REGION Network 13: IW824 - Spare Input
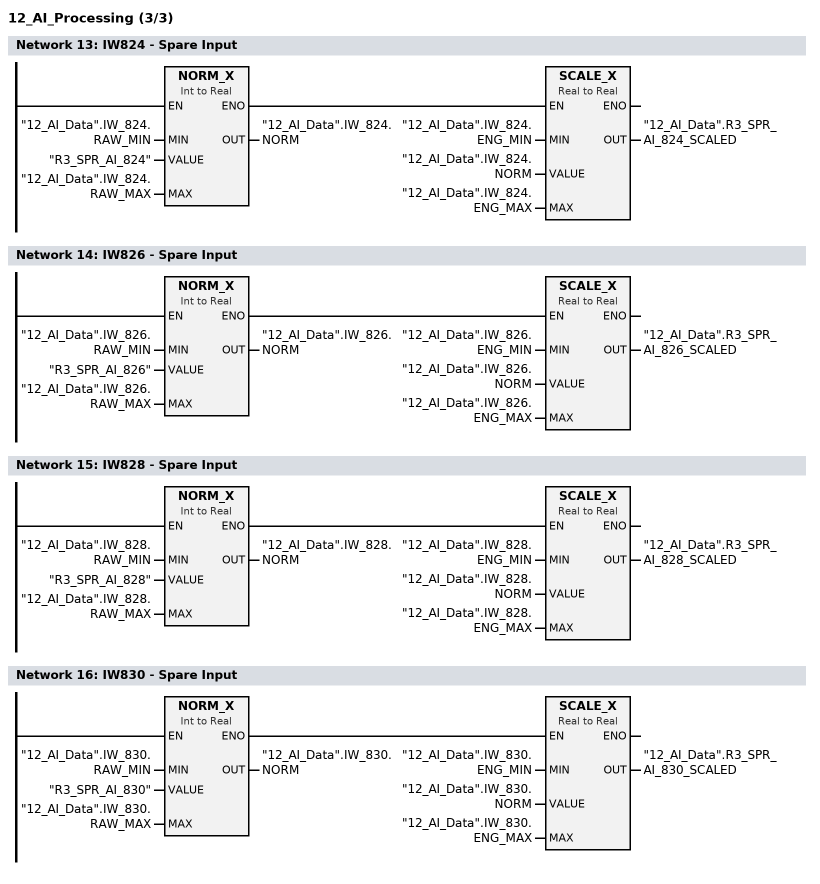
   RUNG wire#powerrail
      { S7_Templates := "[SrcType := Int, DestType := Real]" } Normalize(min := "12_AI_Data".IW_824.RAW_MIN, value := "R3_SPR_AI_824", max := "12_AI_Data".IW_824.RAW_MAX, out => "12_AI_Data".IW_824.NORM)
      { S7_Templates := "[SrcType := Real, DestType := Real]" } Scale(min := "12_AI_Data".IW_824.ENG_MIN, value := "12_AI_Data".IW_824.NORM, max := "12_AI_Data".IW_824.ENG_MAX, out => "12_AI_Data".R3_SPR_AI_824_SCALED)
   END_RUNG
   // the same network as SCL:
   "12_AI_Data".IW_824.NORM := NORM_X(MIN := "12_AI_Data".IW_824.RAW_MIN, VALUE := "R3_SPR_AI_824", MAX := "12_AI_Data".IW_824.RAW_MAX);
   "12_AI_Data".R3_SPR_AI_824_SCALED := SCALE_X(MIN := "12_AI_Data".IW_824.ENG_MIN, VALUE := "12_AI_Data".IW_824.NORM, MAX := "12_AI_Data".IW_824.ENG_MAX);
END_REGION

REGION Network 14: IW826 - Spare Input
   RUNG wire#powerrail
      { S7_Templates := "[SrcType := Int, DestType := Real]" } Normalize(min := "12_AI_Data".IW_826.RAW_MIN, value := "R3_SPR_AI_826", max := "12_AI_Data".IW_826.RAW_MAX, out => "12_AI_Data".IW_826.NORM)
      { S7_Templates := "[SrcType := Real, DestType := Real]" } Scale(min := "12_AI_Data".IW_826.ENG_MIN, value := "12_AI_Data".IW_826.NORM, max := "12_AI_Data".IW_826.ENG_MAX, out => "12_AI_Data".R3_SPR_AI_826_SCALED)
   END_RUNG
   // the same network as SCL:
   "12_AI_Data".IW_826.NORM := NORM_X(MIN := "12_AI_Data".IW_826.RAW_MIN, VALUE := "R3_SPR_AI_826", MAX := "12_AI_Data".IW_826.RAW_MAX);
   "12_AI_Data".R3_SPR_AI_826_SCALED := SCALE_X(MIN := "12_AI_Data".IW_826.ENG_MIN, VALUE := "12_AI_Data".IW_826.NORM, MAX := "12_AI_Data".IW_826.ENG_MAX);
END_REGION

REGION Network 15: IW828 - Spare Input
   RUNG wire#powerrail
      { S7_Templates := "[SrcType := Int, DestType := Real]" } Normalize(min := "12_AI_Data".IW_828.RAW_MIN, value := "R3_SPR_AI_828", max := "12_AI_Data".IW_828.RAW_MAX, out => "12_AI_Data".IW_828.NORM)
      { S7_Templates := "[SrcType := Real, DestType := Real]" } Scale(min := "12_AI_Data".IW_828.ENG_MIN, value := "12_AI_Data".IW_828.NORM, max := "12_AI_Data".IW_828.ENG_MAX, out => "12_AI_Data".R3_SPR_AI_828_SCALED)
   END_RUNG
   // the same network as SCL:
   "12_AI_Data".IW_828.NORM := NORM_X(MIN := "12_AI_Data".IW_828.RAW_MIN, VALUE := "R3_SPR_AI_828", MAX := "12_AI_Data".IW_828.RAW_MAX);
   "12_AI_Data".R3_SPR_AI_828_SCALED := SCALE_X(MIN := "12_AI_Data".IW_828.ENG_MIN, VALUE := "12_AI_Data".IW_828.NORM, MAX := "12_AI_Data".IW_828.ENG_MAX);
END_REGION

REGION Network 16: IW830 - Spare Input
   RUNG wire#powerrail
      { S7_Templates := "[SrcType := Int, DestType := Real]" } Normalize(min := "12_AI_Data".IW_830.RAW_MIN, value := "R3_SPR_AI_830", max := "12_AI_Data".IW_830.RAW_MAX, out => "12_AI_Data".IW_830.NORM)
      { S7_Templates := "[SrcType := Real, DestType := Real]" } Scale(min := "12_AI_Data".IW_830.ENG_MIN, value := "12_AI_Data".IW_830.NORM, max := "12_AI_Data".IW_830.ENG_MAX, out => "12_AI_Data".R3_SPR_AI_830_SCALED)
   END_RUNG
   // the same network as SCL:
   "12_AI_Data".IW_830.NORM := NORM_X(MIN := "12_AI_Data".IW_830.RAW_MIN, VALUE := "R3_SPR_AI_830", MAX := "12_AI_Data".IW_830.RAW_MAX);
   "12_AI_Data".R3_SPR_AI_830_SCALED := SCALE_X(MIN := "12_AI_Data".IW_830.ENG_MIN, VALUE := "12_AI_Data".IW_830.NORM, MAX := "12_AI_Data".IW_830.ENG_MAX);
END_REGION
END_FUNCTION

FUNCTION "14_DQ_Processing" : Void   // FC14, LAD
TITLE = Digital Output Processing
{ S7_Optimized_Access := 'TRUE' }
AUTHOR : JRS
VERSION : 0.1
// To process code outputs prior to physical connection
BEGIN

REGION Network 1: Q136.0 - Fresh Water Fill Valve Control (CV-358)
   // True = OPEN, False = CLOSE
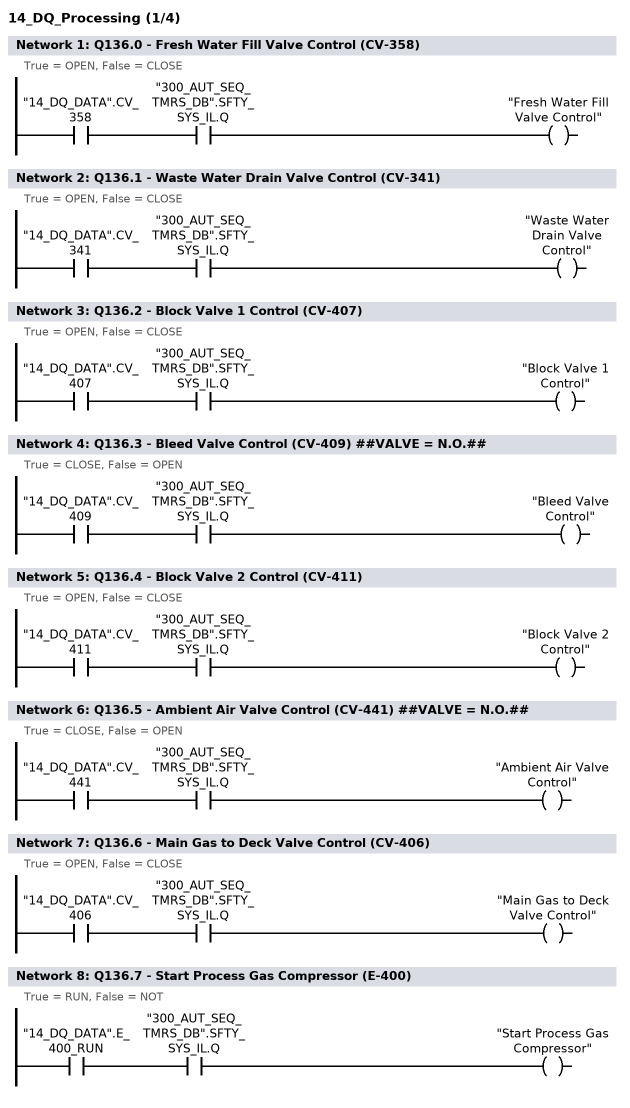
   RUNG wire#powerrail
      Contact( "14_DQ_DATA".CV_358 )
      Contact( "300_AUT_SEQ_TMRS_DB".SFTY_SYS_IL.Q )
      Coil( "Fresh Water Fill Valve Control" )
   END_RUNG
   // the same network as SCL:
   "Fresh Water Fill Valve Control" := "14_DQ_DATA".CV_358 AND "300_AUT_SEQ_TMRS_DB".SFTY_SYS_IL.Q;
END_REGION

REGION Network 2: Q136.1 - Waste Water Drain Valve Control (CV-341)
   // True = OPEN, False = CLOSE
   RUNG wire#powerrail
      Contact( "14_DQ_DATA".CV_341 )
      Contact( "300_AUT_SEQ_TMRS_DB".SFTY_SYS_IL.Q )
      Coil( "Waste Water Drain Valve Control" )
   END_RUNG
   // the same network as SCL:
   "Waste Water Drain Valve Control" := "14_DQ_DATA".CV_341 AND "300_AUT_SEQ_TMRS_DB".SFTY_SYS_IL.Q;
END_REGION

REGION Network 3: Q136.2 - Block Valve 1 Control (CV-407)
   // True = OPEN, False = CLOSE
   RUNG wire#powerrail
      Contact( "14_DQ_DATA".CV_407 )
      Contact( "300_AUT_SEQ_TMRS_DB".SFTY_SYS_IL.Q )
      Coil( "Block Valve 1 Control" )
   END_RUNG
   // the same network as SCL:
   "Block Valve 1 Control" := "14_DQ_DATA".CV_407 AND "300_AUT_SEQ_TMRS_DB".SFTY_SYS_IL.Q;
END_REGION

REGION Network 4: Q136.3 - Bleed Valve Control (CV-409) ##VALVE = N.O.##
   // True = CLOSE, False = OPEN
   RUNG wire#powerrail
      Contact( "14_DQ_DATA".CV_409 )
      Contact( "300_AUT_SEQ_TMRS_DB".SFTY_SYS_IL.Q )
      Coil( "Bleed Valve Control" )
   END_RUNG
   // the same network as SCL:
   "Bleed Valve Control" := "14_DQ_DATA".CV_409 AND "300_AUT_SEQ_TMRS_DB".SFTY_SYS_IL.Q;
END_REGION

REGION Network 5: Q136.4 - Block Valve 2 Control (CV-411)
   // True = OPEN, False = CLOSE
   RUNG wire#powerrail
      Contact( "14_DQ_DATA".CV_411 )
      Contact( "300_AUT_SEQ_TMRS_DB".SFTY_SYS_IL.Q )
      Coil( "Block Valve 2 Control" )
   END_RUNG
   // the same network as SCL:
   "Block Valve 2 Control" := "14_DQ_DATA".CV_411 AND "300_AUT_SEQ_TMRS_DB".SFTY_SYS_IL.Q;
END_REGION

REGION Network 6: Q136.5 - Ambient Air Valve Control (CV-441) ##VALVE = N.O.##
   // True = CLOSE, False = OPEN
   RUNG wire#powerrail
      Contact( "14_DQ_DATA".CV_441 )
      Contact( "300_AUT_SEQ_TMRS_DB".SFTY_SYS_IL.Q )
      Coil( "Ambient Air Valve Control" )
   END_RUNG
   // the same network as SCL:
   "Ambient Air Valve Control" := "14_DQ_DATA".CV_441 AND "300_AUT_SEQ_TMRS_DB".SFTY_SYS_IL.Q;
END_REGION

REGION Network 7: Q136.6 - Main Gas to Deck Valve Control (CV-406)
   // True = OPEN, False = CLOSE
   RUNG wire#powerrail
      Contact( "14_DQ_DATA".CV_406 )
      Contact( "300_AUT_SEQ_TMRS_DB".SFTY_SYS_IL.Q )
      Coil( "Main Gas to Deck Valve Control" )
   END_RUNG
   // the same network as SCL:
   "Main Gas to Deck Valve Control" := "14_DQ_DATA".CV_406 AND "300_AUT_SEQ_TMRS_DB".SFTY_SYS_IL.Q;
END_REGION

REGION Network 8: Q136.7 - Start Process Gas Compressor (E-400)
   // True = RUN, False = NOT
   RUNG wire#powerrail
      Contact( "14_DQ_DATA".E_400_RUN )
      Contact( "300_AUT_SEQ_TMRS_DB".SFTY_SYS_IL.Q )
      Coil( "Start Process Gas Compressor" )
   END_RUNG
   // the same network as SCL:
   "Start Process Gas Compressor" := "14_DQ_DATA".E_400_RUN AND "300_AUT_SEQ_TMRS_DB".SFTY_SYS_IL.Q;
END_REGION

REGION Network 9: Q137.0 - GCU Recirculation Pump Control (P-303)
   // True = RUN, False = NOT
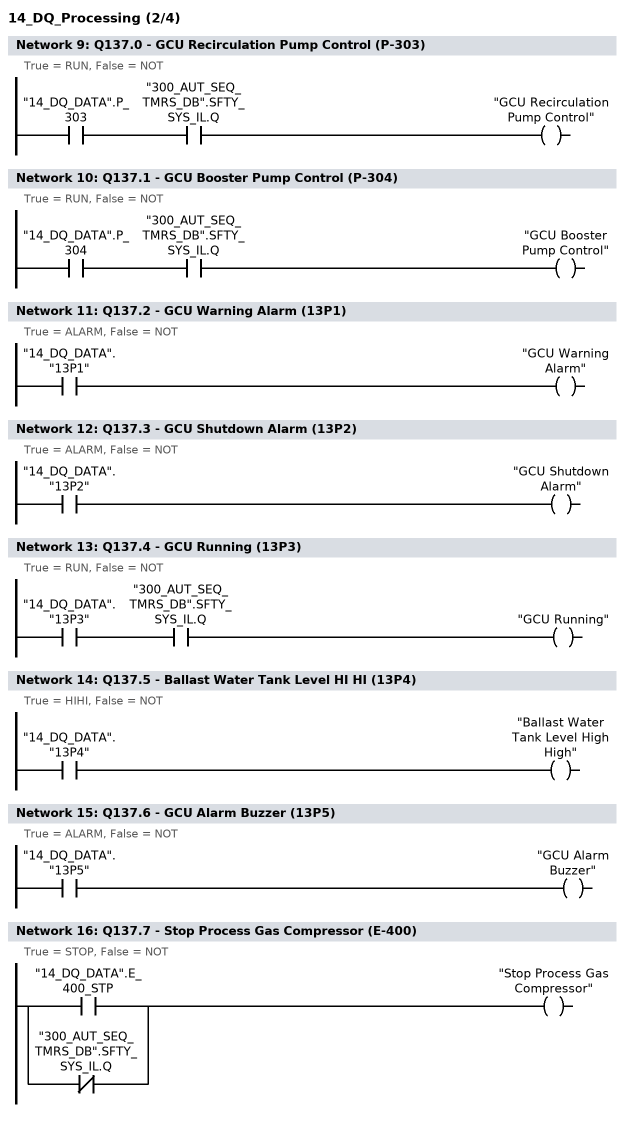
   RUNG wire#powerrail
      Contact( "14_DQ_DATA".P_303 )
      Contact( "300_AUT_SEQ_TMRS_DB".SFTY_SYS_IL.Q )
      Coil( "GCU Recirculation Pump Control" )
   END_RUNG
   // the same network as SCL:
   "GCU Recirculation Pump Control" := "14_DQ_DATA".P_303 AND "300_AUT_SEQ_TMRS_DB".SFTY_SYS_IL.Q;
END_REGION

REGION Network 10: Q137.1 - GCU Booster Pump Control (P-304)
   // True = RUN, False = NOT
   RUNG wire#powerrail
      Contact( "14_DQ_DATA".P_304 )
      Contact( "300_AUT_SEQ_TMRS_DB".SFTY_SYS_IL.Q )
      Coil( "GCU Booster Pump Control" )
   END_RUNG
   // the same network as SCL:
   "GCU Booster Pump Control" := "14_DQ_DATA".P_304 AND "300_AUT_SEQ_TMRS_DB".SFTY_SYS_IL.Q;
END_REGION

REGION Network 11: Q137.2 - GCU Warning Alarm (13P1)
   // True = ALARM, False = NOT
   RUNG wire#powerrail
      Contact( "14_DQ_DATA"."13P1" )
      Coil( "GCU Warning Alarm" )
   END_RUNG
   // the same network as SCL:
   "GCU Warning Alarm" := "14_DQ_DATA"."13P1";
END_REGION

REGION Network 12: Q137.3 - GCU Shutdown Alarm (13P2)
   // True = ALARM, False = NOT
   RUNG wire#powerrail
      Contact( "14_DQ_DATA"."13P2" )
      Coil( "GCU Shutdown Alarm" )
   END_RUNG
   // the same network as SCL:
   "GCU Shutdown Alarm" := "14_DQ_DATA"."13P2";
END_REGION

REGION Network 13: Q137.4 - GCU Running (13P3)
   // True = RUN, False = NOT
   RUNG wire#powerrail
      Contact( "14_DQ_DATA"."13P3" )
      Contact( "300_AUT_SEQ_TMRS_DB".SFTY_SYS_IL.Q )
      Coil( "GCU Running" )
   END_RUNG
   // the same network as SCL:
   "GCU Running" := "14_DQ_DATA"."13P3" AND "300_AUT_SEQ_TMRS_DB".SFTY_SYS_IL.Q;
END_REGION

REGION Network 14: Q137.5 - Ballast Water Tank Level HI HI (13P4)
   // True = HIHI, False = NOT
   RUNG wire#powerrail
      Contact( "14_DQ_DATA"."13P4" )
      Coil( "Ballast Water Tank Level High High" )
   END_RUNG
   // the same network as SCL:
   "Ballast Water Tank Level High High" := "14_DQ_DATA"."13P4";
END_REGION

REGION Network 15: Q137.6 - GCU Alarm Buzzer (13P5)
   // True = ALARM, False = NOT
   RUNG wire#powerrail
      Contact( "14_DQ_DATA"."13P5" )
      Coil( "GCU Alarm Buzzer" )
   END_RUNG
   // the same network as SCL:
   "GCU Alarm Buzzer" := "14_DQ_DATA"."13P5";
END_REGION

REGION Network 16: Q137.7 - Stop Process Gas Compressor (E-400)
   // True = STOP, False = NOT
   RUNG wire#powerrail
      Contact( "14_DQ_DATA".E_400_STP )
      wire#w1
      Coil( "Stop Process Gas Compressor" )
   END_RUNG
   RUNG wire#powerrail
      I_Contact( "300_AUT_SEQ_TMRS_DB".SFTY_SYS_IL.Q )
   END_RUNG wire#w1
   // the same network as SCL:
   "Stop Process Gas Compressor" := "14_DQ_DATA".E_400_STP OR NOT "300_AUT_SEQ_TMRS_DB".SFTY_SYS_IL.Q;
END_REGION

REGION Network 17: Q138.0 - Pilot For GTT FPT Valve (CV-422-FPT)
   // True = OPEN, False = CLOSE
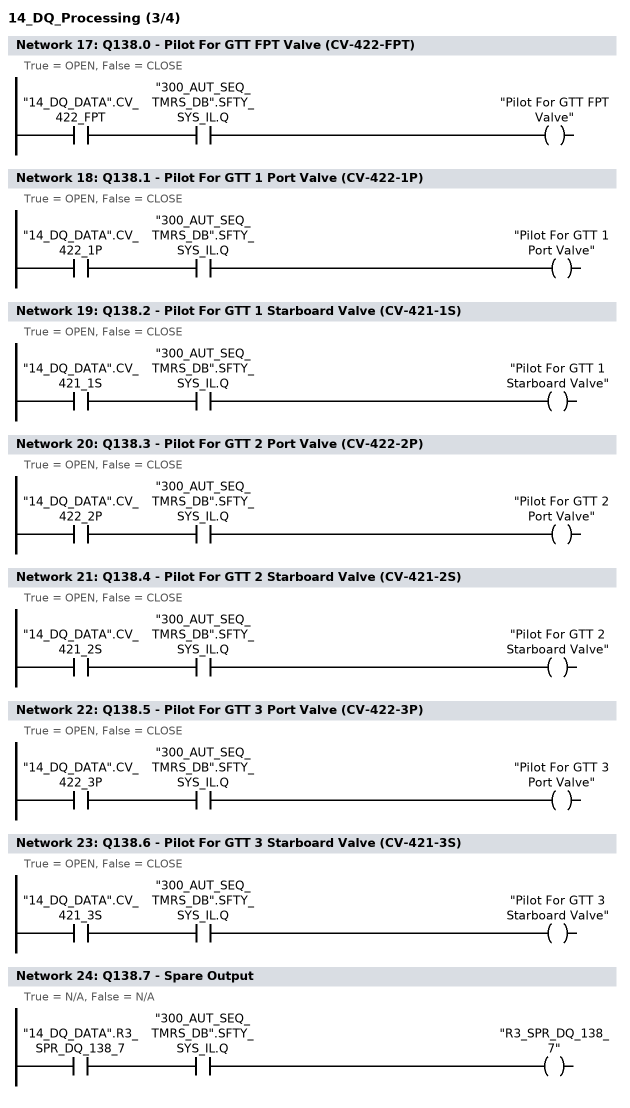
   RUNG wire#powerrail
      Contact( "14_DQ_DATA".CV_422_FPT )
      Contact( "300_AUT_SEQ_TMRS_DB".SFTY_SYS_IL.Q )
      Coil( "Pilot For GTT FPT Valve" )
   END_RUNG
   // the same network as SCL:
   "Pilot For GTT FPT Valve" := "14_DQ_DATA".CV_422_FPT AND "300_AUT_SEQ_TMRS_DB".SFTY_SYS_IL.Q;
END_REGION

REGION Network 18: Q138.1 - Pilot For GTT 1 Port Valve (CV-422-1P)
   // True = OPEN, False = CLOSE
   RUNG wire#powerrail
      Contact( "14_DQ_DATA".CV_422_1P )
      Contact( "300_AUT_SEQ_TMRS_DB".SFTY_SYS_IL.Q )
      Coil( "Pilot For GTT 1 Port Valve" )
   END_RUNG
   // the same network as SCL:
   "Pilot For GTT 1 Port Valve" := "14_DQ_DATA".CV_422_1P AND "300_AUT_SEQ_TMRS_DB".SFTY_SYS_IL.Q;
END_REGION

REGION Network 19: Q138.2 - Pilot For GTT 1 Starboard Valve (CV-421-1S)
   // True = OPEN, False = CLOSE
   RUNG wire#powerrail
      Contact( "14_DQ_DATA".CV_421_1S )
      Contact( "300_AUT_SEQ_TMRS_DB".SFTY_SYS_IL.Q )
      Coil( "Pilot For GTT 1 Starboard Valve" )
   END_RUNG
   // the same network as SCL:
   "Pilot For GTT 1 Starboard Valve" := "14_DQ_DATA".CV_421_1S AND "300_AUT_SEQ_TMRS_DB".SFTY_SYS_IL.Q;
END_REGION

REGION Network 20: Q138.3 - Pilot For GTT 2 Port Valve (CV-422-2P)
   // True = OPEN, False = CLOSE
   RUNG wire#powerrail
      Contact( "14_DQ_DATA".CV_422_2P )
      Contact( "300_AUT_SEQ_TMRS_DB".SFTY_SYS_IL.Q )
      Coil( "Pilot For GTT 2 Port Valve" )
   END_RUNG
   // the same network as SCL:
   "Pilot For GTT 2 Port Valve" := "14_DQ_DATA".CV_422_2P AND "300_AUT_SEQ_TMRS_DB".SFTY_SYS_IL.Q;
END_REGION

REGION Network 21: Q138.4 - Pilot For GTT 2 Starboard Valve (CV-421-2S)
   // True = OPEN, False = CLOSE
   RUNG wire#powerrail
      Contact( "14_DQ_DATA".CV_421_2S )
      Contact( "300_AUT_SEQ_TMRS_DB".SFTY_SYS_IL.Q )
      Coil( "Pilot For GTT 2 Starboard Valve" )
   END_RUNG
   // the same network as SCL:
   "Pilot For GTT 2 Starboard Valve" := "14_DQ_DATA".CV_421_2S AND "300_AUT_SEQ_TMRS_DB".SFTY_SYS_IL.Q;
END_REGION

REGION Network 22: Q138.5 - Pilot For GTT 3 Port Valve (CV-422-3P)
   // True = OPEN, False = CLOSE
   RUNG wire#powerrail
      Contact( "14_DQ_DATA".CV_422_3P )
      Contact( "300_AUT_SEQ_TMRS_DB".SFTY_SYS_IL.Q )
      Coil( "Pilot For GTT 3 Port Valve" )
   END_RUNG
   // the same network as SCL:
   "Pilot For GTT 3 Port Valve" := "14_DQ_DATA".CV_422_3P AND "300_AUT_SEQ_TMRS_DB".SFTY_SYS_IL.Q;
END_REGION

REGION Network 23: Q138.6 - Pilot For GTT 3 Starboard Valve (CV-421-3S)
   // True = OPEN, False = CLOSE
   RUNG wire#powerrail
      Contact( "14_DQ_DATA".CV_421_3S )
      Contact( "300_AUT_SEQ_TMRS_DB".SFTY_SYS_IL.Q )
      Coil( "Pilot For GTT 3 Starboard Valve" )
   END_RUNG
   // the same network as SCL:
   "Pilot For GTT 3 Starboard Valve" := "14_DQ_DATA".CV_421_3S AND "300_AUT_SEQ_TMRS_DB".SFTY_SYS_IL.Q;
END_REGION

REGION Network 24: Q138.7 - Spare Output
   // True = N/A, False = N/A
   RUNG wire#powerrail
      Contact( "14_DQ_DATA".R3_SPR_DQ_138_7 )
      Contact( "300_AUT_SEQ_TMRS_DB".SFTY_SYS_IL.Q )
      Coil( "R3_SPR_DQ_138_7" )
   END_RUNG
   // the same network as SCL:
   "R3_SPR_DQ_138_7" := "14_DQ_DATA".R3_SPR_DQ_138_7 AND "300_AUT_SEQ_TMRS_DB".SFTY_SYS_IL.Q;
END_REGION

REGION Network 25: Q139.0 - Pilot For GTT 4 Port Valve (CV-422-4P)
   // True = OPEN, False = CLOSE
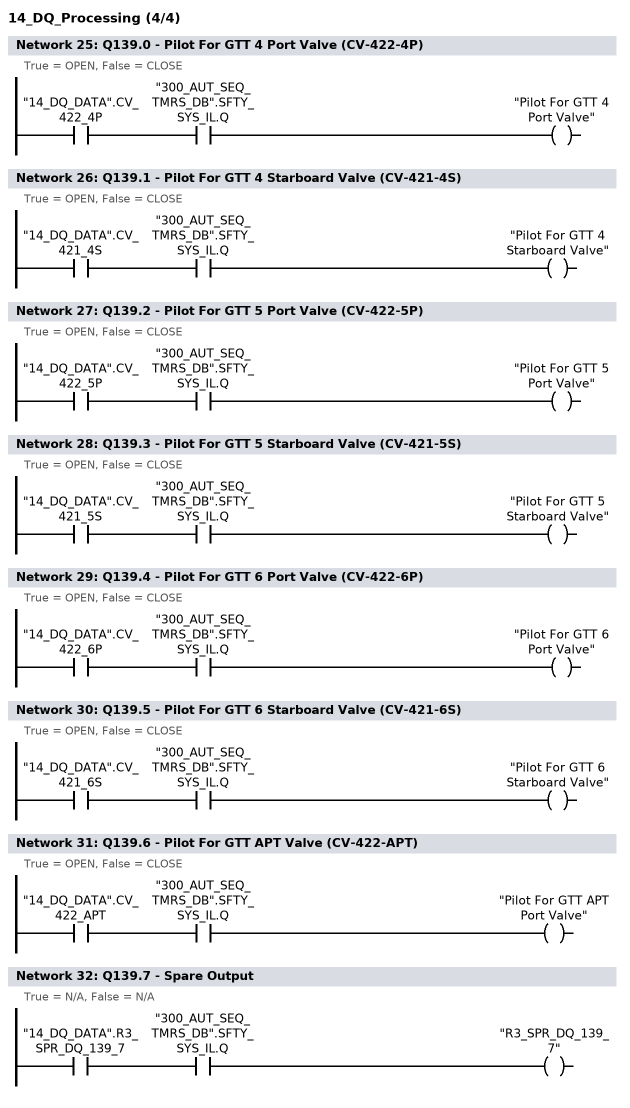
   RUNG wire#powerrail
      Contact( "14_DQ_DATA".CV_422_4P )
      Contact( "300_AUT_SEQ_TMRS_DB".SFTY_SYS_IL.Q )
      Coil( "Pilot For GTT 4 Port Valve" )
   END_RUNG
   // the same network as SCL:
   "Pilot For GTT 4 Port Valve" := "14_DQ_DATA".CV_422_4P AND "300_AUT_SEQ_TMRS_DB".SFTY_SYS_IL.Q;
END_REGION

REGION Network 26: Q139.1 - Pilot For GTT 4 Starboard Valve (CV-421-4S)
   // True = OPEN, False = CLOSE
   RUNG wire#powerrail
      Contact( "14_DQ_DATA".CV_421_4S )
      Contact( "300_AUT_SEQ_TMRS_DB".SFTY_SYS_IL.Q )
      Coil( "Pilot For GTT 4 Starboard Valve" )
   END_RUNG
   // the same network as SCL:
   "Pilot For GTT 4 Starboard Valve" := "14_DQ_DATA".CV_421_4S AND "300_AUT_SEQ_TMRS_DB".SFTY_SYS_IL.Q;
END_REGION

REGION Network 27: Q139.2 - Pilot For GTT 5 Port Valve (CV-422-5P)
   // True = OPEN, False = CLOSE
   RUNG wire#powerrail
      Contact( "14_DQ_DATA".CV_422_5P )
      Contact( "300_AUT_SEQ_TMRS_DB".SFTY_SYS_IL.Q )
      Coil( "Pilot For GTT 5 Port Valve" )
   END_RUNG
   // the same network as SCL:
   "Pilot For GTT 5 Port Valve" := "14_DQ_DATA".CV_422_5P AND "300_AUT_SEQ_TMRS_DB".SFTY_SYS_IL.Q;
END_REGION

REGION Network 28: Q139.3 - Pilot For GTT 5 Starboard Valve (CV-421-5S)
   // True = OPEN, False = CLOSE
   RUNG wire#powerrail
      Contact( "14_DQ_DATA".CV_421_5S )
      Contact( "300_AUT_SEQ_TMRS_DB".SFTY_SYS_IL.Q )
      Coil( "Pilot For GTT 5 Starboard Valve" )
   END_RUNG
   // the same network as SCL:
   "Pilot For GTT 5 Starboard Valve" := "14_DQ_DATA".CV_421_5S AND "300_AUT_SEQ_TMRS_DB".SFTY_SYS_IL.Q;
END_REGION

REGION Network 29: Q139.4 - Pilot For GTT 6 Port Valve (CV-422-6P)
   // True = OPEN, False = CLOSE
   RUNG wire#powerrail
      Contact( "14_DQ_DATA".CV_422_6P )
      Contact( "300_AUT_SEQ_TMRS_DB".SFTY_SYS_IL.Q )
      Coil( "Pilot For GTT 6 Port Valve" )
   END_RUNG
   // the same network as SCL:
   "Pilot For GTT 6 Port Valve" := "14_DQ_DATA".CV_422_6P AND "300_AUT_SEQ_TMRS_DB".SFTY_SYS_IL.Q;
END_REGION

REGION Network 30: Q139.5 - Pilot For GTT 6 Starboard Valve (CV-421-6S)
   // True = OPEN, False = CLOSE
   RUNG wire#powerrail
      Contact( "14_DQ_DATA".CV_421_6S )
      Contact( "300_AUT_SEQ_TMRS_DB".SFTY_SYS_IL.Q )
      Coil( "Pilot For GTT 6 Starboard Valve" )
   END_RUNG
   // the same network as SCL:
   "Pilot For GTT 6 Starboard Valve" := "14_DQ_DATA".CV_421_6S AND "300_AUT_SEQ_TMRS_DB".SFTY_SYS_IL.Q;
END_REGION

REGION Network 31: Q139.6 - Pilot For GTT APT Valve (CV-422-APT)
   // True = OPEN, False = CLOSE
   RUNG wire#powerrail
      Contact( "14_DQ_DATA".CV_422_APT )
      Contact( "300_AUT_SEQ_TMRS_DB".SFTY_SYS_IL.Q )
      Coil( "Pilot For GTT APT Port Valve" )
   END_RUNG
   // the same network as SCL:
   "Pilot For GTT APT Port Valve" := "14_DQ_DATA".CV_422_APT AND "300_AUT_SEQ_TMRS_DB".SFTY_SYS_IL.Q;
END_REGION

REGION Network 32: Q139.7 - Spare Output
   // True = N/A, False = N/A
   RUNG wire#powerrail
      Contact( "14_DQ_DATA".R3_SPR_DQ_139_7 )
      Contact( "300_AUT_SEQ_TMRS_DB".SFTY_SYS_IL.Q )
      Coil( "R3_SPR_DQ_139_7" )
   END_RUNG
   // the same network as SCL:
   "R3_SPR_DQ_139_7" := "14_DQ_DATA".R3_SPR_DQ_139_7 AND "300_AUT_SEQ_TMRS_DB".SFTY_SYS_IL.Q;
END_REGION
END_FUNCTION

FUNCTION "16_AQ_Processing" : Void   // FC16, LAD
TITLE = Analogue Output Processing
{ S7_Optimized_Access := 'TRUE' }
AUTHOR : JRS
VERSION : 0.1
// To process code outputs prior to physical connection
BEGIN

REGION Network 1: QW800 - Gas Vent Position Control (CV-405)
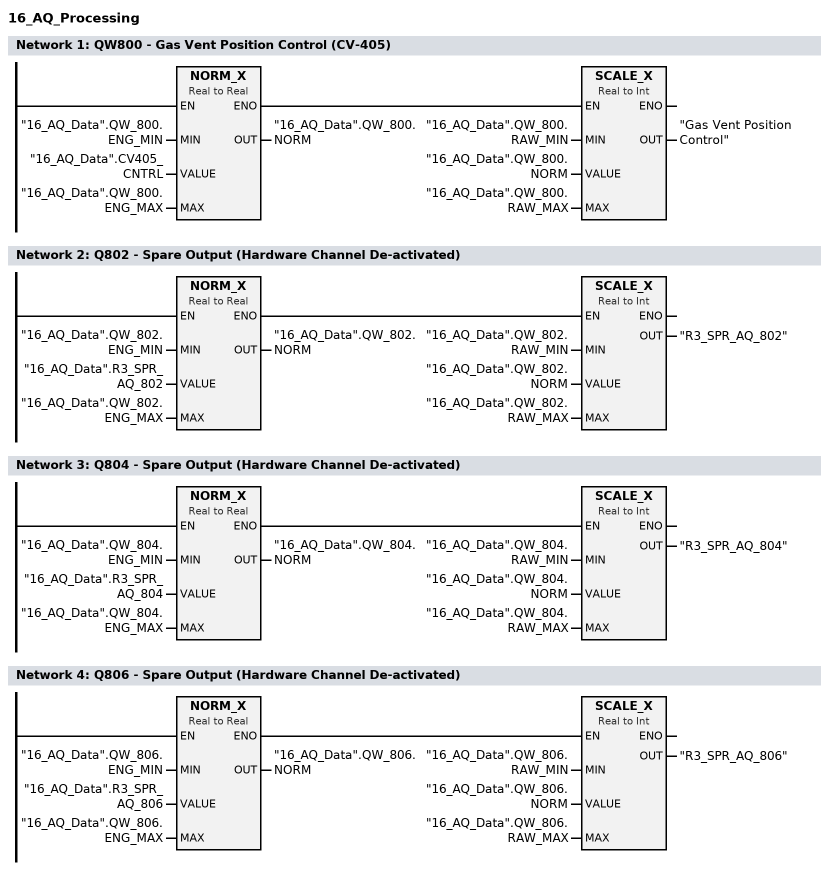
   RUNG wire#powerrail
      { S7_Templates := "[SrcType := Real, DestType := Real]" } Normalize(min := "16_AQ_Data".QW_800.ENG_MIN, value := "16_AQ_Data".CV405_CNTRL, max := "16_AQ_Data".QW_800.ENG_MAX, out => "16_AQ_Data".QW_800.NORM)
      { S7_Templates := "[SrcType := Real, DestType := Int]" } Scale(min := "16_AQ_Data".QW_800.RAW_MIN, value := "16_AQ_Data".QW_800.NORM, max := "16_AQ_Data".QW_800.RAW_MAX, out => "Gas Vent Position Control")
   END_RUNG
   // the same network as SCL:
   "16_AQ_Data".QW_800.NORM := NORM_X(MIN := "16_AQ_Data".QW_800.ENG_MIN, VALUE := "16_AQ_Data".CV405_CNTRL, MAX := "16_AQ_Data".QW_800.ENG_MAX);
   "Gas Vent Position Control" := SCALE_X(MIN := "16_AQ_Data".QW_800.RAW_MIN, VALUE := "16_AQ_Data".QW_800.NORM, MAX := "16_AQ_Data".QW_800.RAW_MAX);
END_REGION

REGION Network 2: Q802 - Spare Output (Hardware Channel De-activated)
   RUNG wire#powerrail
      { S7_Templates := "[SrcType := Real, DestType := Real]" } Normalize(min := "16_AQ_Data".QW_802.ENG_MIN, value := "16_AQ_Data".R3_SPR_AQ_802, max := "16_AQ_Data".QW_802.ENG_MAX, out => "16_AQ_Data".QW_802.NORM)
      { S7_Templates := "[SrcType := Real, DestType := Int]" } Scale(min := "16_AQ_Data".QW_802.RAW_MIN, value := "16_AQ_Data".QW_802.NORM, max := "16_AQ_Data".QW_802.RAW_MAX, out => "R3_SPR_AQ_802")
   END_RUNG
   // the same network as SCL:
   "16_AQ_Data".QW_802.NORM := NORM_X(MIN := "16_AQ_Data".QW_802.ENG_MIN, VALUE := "16_AQ_Data".R3_SPR_AQ_802, MAX := "16_AQ_Data".QW_802.ENG_MAX);
   "R3_SPR_AQ_802" := SCALE_X(MIN := "16_AQ_Data".QW_802.RAW_MIN, VALUE := "16_AQ_Data".QW_802.NORM, MAX := "16_AQ_Data".QW_802.RAW_MAX);
END_REGION

REGION Network 3: Q804 - Spare Output (Hardware Channel De-activated)
   RUNG wire#powerrail
      { S7_Templates := "[SrcType := Real, DestType := Real]" } Normalize(min := "16_AQ_Data".QW_804.ENG_MIN, value := "16_AQ_Data".R3_SPR_AQ_804, max := "16_AQ_Data".QW_804.ENG_MAX, out => "16_AQ_Data".QW_804.NORM)
      { S7_Templates := "[SrcType := Real, DestType := Int]" } Scale(min := "16_AQ_Data".QW_804.RAW_MIN, value := "16_AQ_Data".QW_804.NORM, max := "16_AQ_Data".QW_804.RAW_MAX, out => "R3_SPR_AQ_804")
   END_RUNG
   // the same network as SCL:
   "16_AQ_Data".QW_804.NORM := NORM_X(MIN := "16_AQ_Data".QW_804.ENG_MIN, VALUE := "16_AQ_Data".R3_SPR_AQ_804, MAX := "16_AQ_Data".QW_804.ENG_MAX);
   "R3_SPR_AQ_804" := SCALE_X(MIN := "16_AQ_Data".QW_804.RAW_MIN, VALUE := "16_AQ_Data".QW_804.NORM, MAX := "16_AQ_Data".QW_804.RAW_MAX);
END_REGION

REGION Network 4: Q806 - Spare Output (Hardware Channel De-activated)
   RUNG wire#powerrail
      { S7_Templates := "[SrcType := Real, DestType := Real]" } Normalize(min := "16_AQ_Data".QW_806.ENG_MIN, value := "16_AQ_Data".R3_SPR_AQ_806, max := "16_AQ_Data".QW_806.ENG_MAX, out => "16_AQ_Data".QW_806.NORM)
      { S7_Templates := "[SrcType := Real, DestType := Int]" } Scale(min := "16_AQ_Data".QW_806.RAW_MIN, value := "16_AQ_Data".QW_806.NORM, max := "16_AQ_Data".QW_806.RAW_MAX, out => "R3_SPR_AQ_806")
   END_RUNG
   // the same network as SCL:
   "16_AQ_Data".QW_806.NORM := NORM_X(MIN := "16_AQ_Data".QW_806.ENG_MIN, VALUE := "16_AQ_Data".R3_SPR_AQ_806, MAX := "16_AQ_Data".QW_806.ENG_MAX);
   "R3_SPR_AQ_806" := SCALE_X(MIN := "16_AQ_Data".QW_806.RAW_MIN, VALUE := "16_AQ_Data".QW_806.NORM, MAX := "16_AQ_Data".QW_806.RAW_MAX);
END_REGION
END_FUNCTION

FUNCTION "19_AUTO_CMNDS" : Void   // FC19, LAD
TITLE = Automatic Output Commands
{ S7_Optimized_Access := 'TRUE' }
AUTHOR : JRS
VERSION : 0.1
// To process automatic output commands prior to output processing
   VAR_TEMP   // added for the SCL form of the ladder/FBD networks
      _w1 : Bool;
      _w2 : Bool;
      _w3 : Bool;
      _w4 : Bool;
      _w5 : Bool;
   END_VAR
BEGIN

REGION Network 1: BWTS or BTCS Control (Ballast Water Treatment or Barge Tank Control)
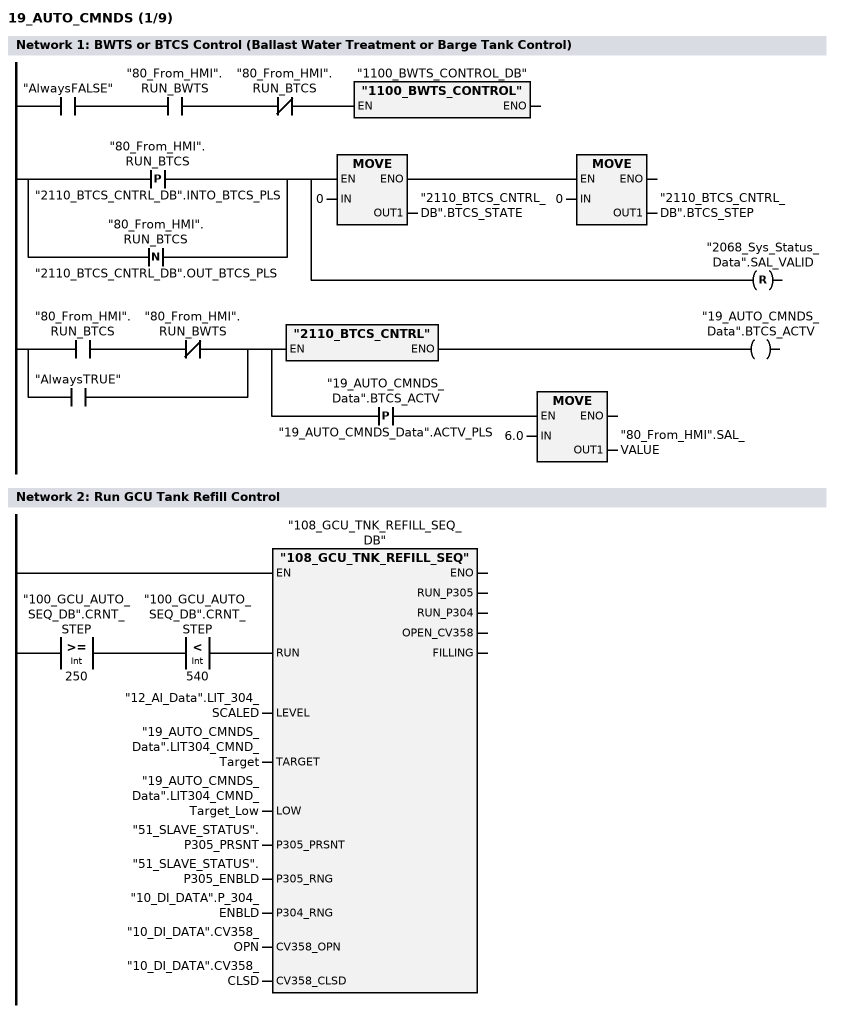
   RUNG wire#powerrail
      Contact( "AlwaysFALSE" )
      Contact( "80_From_HMI".RUN_BWTS )
      I_Contact( "80_From_HMI".RUN_BTCS )
      "1100_BWTS_CONTROL_DB"()
   END_RUNG
   RUNG wire#powerrail
      P_Contact(operand := "80_From_HMI".RUN_BTCS, bit := "2110_BTCS_CNTRL_DB".INTO_BTCS_PLS)
      wire#w1
      Move(in := 0, out1 => "2110_BTCS_CNTRL_DB".BTCS_STATE)
      Move(in := 0, out1 => "2110_BTCS_CNTRL_DB".BTCS_STEP)
   END_RUNG
   RUNG wire#powerrail
      N_Contact(operand := "80_From_HMI".RUN_BTCS, bit := "2110_BTCS_CNTRL_DB".OUT_BTCS_PLS)
   END_RUNG wire#w1
   RUNG wire#w1
      R_Coil( "2068_Sys_Status_Data".SAL_VALID )
   END_RUNG
   RUNG wire#powerrail
      Contact( "80_From_HMI".RUN_BTCS )
      I_Contact( "80_From_HMI".RUN_BWTS )
      wire#w2
      "2110_BTCS_CNTRL"()
      Coil( "19_AUTO_CMNDS_Data".BTCS_ACTV )
   END_RUNG
   RUNG wire#powerrail
      Contact( "AlwaysTRUE" )
   END_RUNG wire#w2
   RUNG wire#w2
      P_Contact(operand := "19_AUTO_CMNDS_Data".BTCS_ACTV, bit := "19_AUTO_CMNDS_Data".ACTV_PLS)
      Move(in := 6.0, out1 => "80_From_HMI".SAL_VALUE)
   END_RUNG
   // the same network as SCL:
   IF "AlwaysFALSE" AND "80_From_HMI".RUN_BWTS AND NOT "80_From_HMI".RUN_BTCS THEN
       "1100_BWTS_CONTROL_DB"();   // "1100_BWTS_CONTROL"
   END_IF;
   #_w1 := "80_From_HMI".RUN_BTCS AND NOT "2110_BTCS_CNTRL_DB".INTO_BTCS_PLS;   // rising edge of "80_From_HMI".RUN_BTCS
   "2110_BTCS_CNTRL_DB".INTO_BTCS_PLS := "80_From_HMI".RUN_BTCS;
   #_w2 := NOT "80_From_HMI".RUN_BTCS AND "2110_BTCS_CNTRL_DB".OUT_BTCS_PLS;   // falling edge of "80_From_HMI".RUN_BTCS
   "2110_BTCS_CNTRL_DB".OUT_BTCS_PLS := "80_From_HMI".RUN_BTCS;
   IF #_w1 OR #_w2 THEN
       "2110_BTCS_CNTRL_DB".BTCS_STATE := 0;
       "2110_BTCS_CNTRL_DB".BTCS_STEP := 0;
       "2068_Sys_Status_Data".SAL_VALID := FALSE;
   END_IF;
   #_w3 := ("80_From_HMI".RUN_BTCS AND NOT "80_From_HMI".RUN_BWTS) OR "AlwaysTRUE";
   "2110_BTCS_CNTRL"(EN := #_w3, ENO => #_w4);
   "19_AUTO_CMNDS_Data".BTCS_ACTV := #_w4;
   #_w5 := #_w3 AND "19_AUTO_CMNDS_Data".BTCS_ACTV AND NOT "19_AUTO_CMNDS_Data".ACTV_PLS;   // rising edge of "19_AUTO_CMNDS_Data".BTCS_ACTV
   "19_AUTO_CMNDS_Data".ACTV_PLS := "19_AUTO_CMNDS_Data".BTCS_ACTV;
   IF #_w5 THEN "80_From_HMI".SAL_VALUE := 6.0; END_IF;
END_REGION

REGION Network 2: Run GCU Tank Refill Control
   RUNG wire#powerrail
      "108_GCU_TNK_REFILL_SEQ_DB"(RUN := wire#w1, LEVEL := "12_AI_Data".LIT_304_SCALED, TARGET := "19_AUTO_CMNDS_Data".LIT304_CMND_Target, LOW := "19_AUTO_CMNDS_Data".LIT304_CMND_Target_Low, P305_PRSNT := "51_SLAVE_STATUS".P305_PRSNT, P305_RNG := "51_SLAVE_STATUS".P305_ENBLD, P304_RNG := "10_DI_DATA".P_304_ENBLD, CV358_OPN := "10_DI_DATA".CV358_OPN, CV358_CLSD := "10_DI_DATA".CV358_CLSD, RUN_P305 =>, RUN_P304 =>, OPEN_CV358 =>, FILLING =>)
   END_RUNG
   RUNG wire#powerrail
      { S7_Templates := "SrcType := Int" } GE_Contact(in1 := "100_GCU_AUTO_SEQ_DB".CRNT_STEP, in2 := 250)
      { S7_Templates := "SrcType := Int" } LT_Contact(in1 := "100_GCU_AUTO_SEQ_DB".CRNT_STEP, in2 := 540)
   END_RUNG wire#w1
   // the same network as SCL:
   "108_GCU_TNK_REFILL_SEQ_DB"(RUN := ("100_GCU_AUTO_SEQ_DB".CRNT_STEP >= 250) AND ("100_GCU_AUTO_SEQ_DB".CRNT_STEP < 540),   // "108_GCU_TNK_REFILL_SEQ"
                           LEVEL := "12_AI_Data".LIT_304_SCALED,
                           TARGET := "19_AUTO_CMNDS_Data".LIT304_CMND_Target,
                           LOW := "19_AUTO_CMNDS_Data".LIT304_CMND_Target_Low,
                           P305_PRSNT := "51_SLAVE_STATUS".P305_PRSNT,
                           P305_RNG := "51_SLAVE_STATUS".P305_ENBLD,
                           P304_RNG := "10_DI_DATA".P_304_ENBLD,
                           CV358_OPN := "10_DI_DATA".CV358_OPN,
                           CV358_CLSD := "10_DI_DATA".CV358_CLSD);
END_REGION

REGION Network 3: Run GCU Tank Flush Control
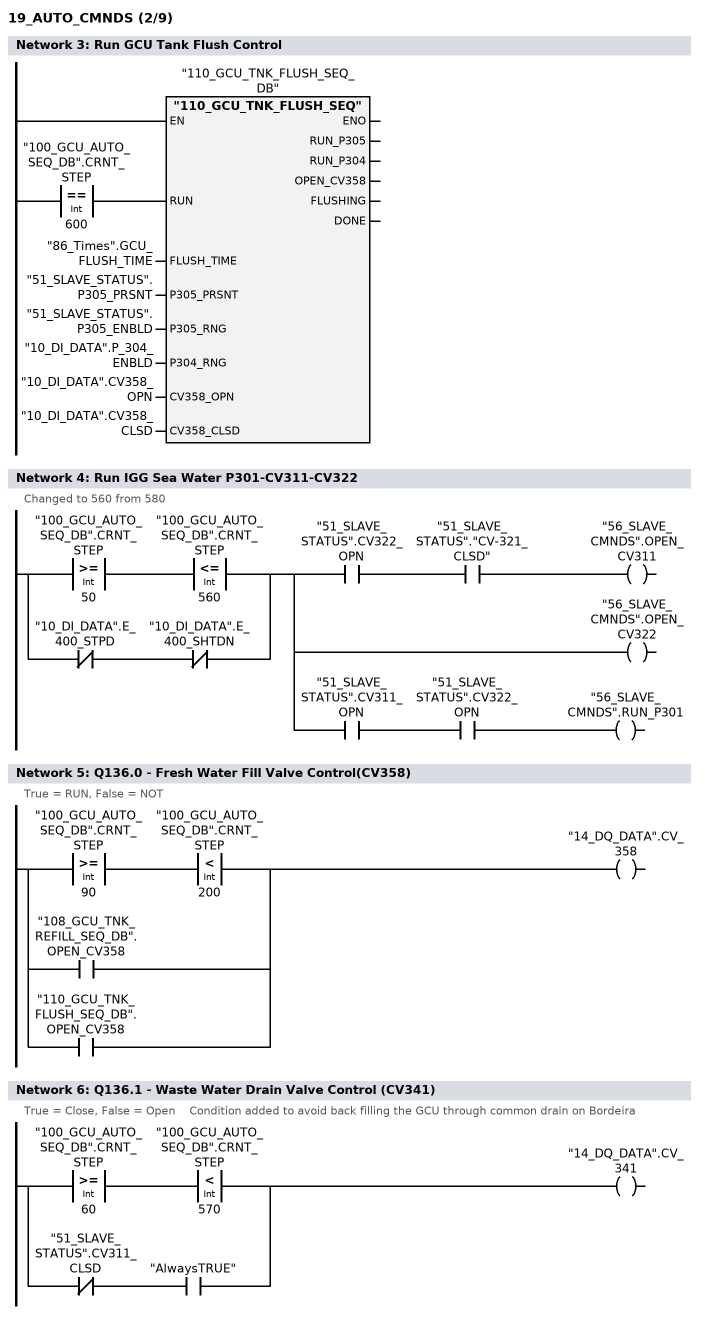
   RUNG wire#powerrail
      "110_GCU_TNK_FLUSH_SEQ_DB"(RUN := wire#w1, FLUSH_TIME := "86_Times".GCU_FLUSH_TIME, P305_PRSNT := "51_SLAVE_STATUS".P305_PRSNT, P305_RNG := "51_SLAVE_STATUS".P305_ENBLD, P304_RNG := "10_DI_DATA".P_304_ENBLD, CV358_OPN := "10_DI_DATA".CV358_OPN, CV358_CLSD := "10_DI_DATA".CV358_CLSD, RUN_P305 =>, RUN_P304 =>, OPEN_CV358 =>, FLUSHING =>, DONE =>)
   END_RUNG
   RUNG wire#powerrail
      { S7_Templates := "SrcType := Int" } EQ_Contact(in1 := "100_GCU_AUTO_SEQ_DB".CRNT_STEP, in2 := 600)
   END_RUNG wire#w1
   // the same network as SCL:
   "110_GCU_TNK_FLUSH_SEQ_DB"(RUN := "100_GCU_AUTO_SEQ_DB".CRNT_STEP = 600,   // "110_GCU_TNK_FLUSH_SEQ"
                           FLUSH_TIME := "86_Times".GCU_FLUSH_TIME,
                           P305_PRSNT := "51_SLAVE_STATUS".P305_PRSNT,
                           P305_RNG := "51_SLAVE_STATUS".P305_ENBLD,
                           P304_RNG := "10_DI_DATA".P_304_ENBLD,
                           CV358_OPN := "10_DI_DATA".CV358_OPN,
                           CV358_CLSD := "10_DI_DATA".CV358_CLSD);
END_REGION
